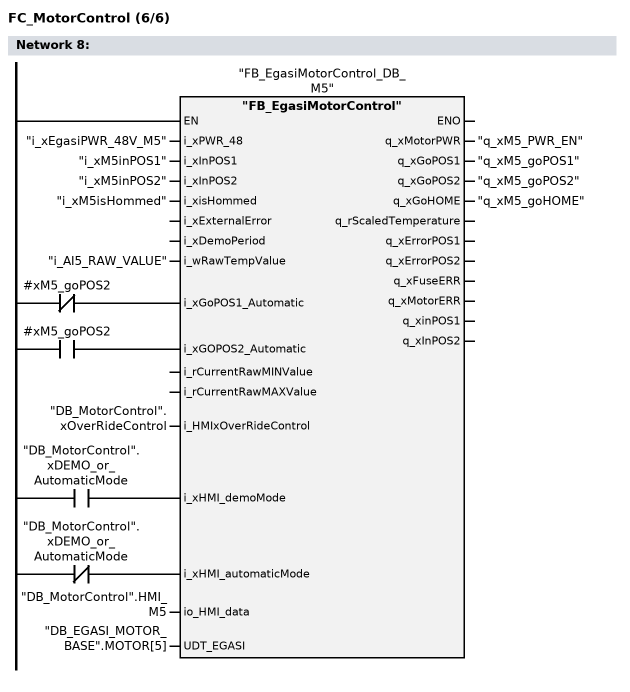
   RUNG wire#powerrail
      "FB_EgasiMotorControl_DB_M5"(i_xGoPOS1_Automatic := wire#w1, i_xGOPOS2_Automatic := wire#w2, i_xHMI_demoMode := wire#w3, i_xHMI_automaticMode := wire#w4, i_xPWR_48 := "i_xEgasiPWR_48V_M5", i_xInPOS1 := "i_xM5inPOS1", i_xInPOS2 := "i_xM5inPOS2", i_xisHommed := "i_xM5isHommed", i_xExternalError :=, i_xDemoPeriod :=, i_wRawTempValue := "i_AI5_RAW_VALUE", i_rCurrentRawMINValue :=, i_rCurrentRawMAXValue :=, i_HMIxOverRideControl := "DB_MotorControl".xOverRideControl, io_HMI_data := "DB_MotorControl".HMI_M5, UDT_EGASI := "DB_EGASI_MOTOR_BASE".MOTOR[5], q_xMotorPWR => "q_xM5_PWR_EN", q_xGoPOS1 => "q_xM5_goPOS1", q_xGoPOS2 => "q_xM5_goPOS2", q_xGoHOME => "q_xM5_goHOME", q_rScaledTemperature =>, q_xErrorPOS1 =>, q_xErrorPOS2 =>, q_xFuseERR =>, q_xMotorERR =>, q_xinPOS1 =>, q_xInPOS2 =>)
   END_RUNG
   RUNG wire#powerrail
      I_Contact( #xM5_goPOS2 )
   END_RUNG wire#w1
   RUNG wire#powerrail
      Contact( #xM5_goPOS2 )
   END_RUNG wire#w2
   RUNG wire#powerrail
      Contact( "DB_MotorControl".xDEMO_or_AutomaticMode )
   END_RUNG wire#w3
   RUNG wire#powerrail
      I_Contact( "DB_MotorControl".xDEMO_or_AutomaticMode )
   END_RUNG wire#w4
   // the same network as SCL:
   "FB_EgasiMotorControl_DB_M5"(i_xPWR_48 := "i_xEgasiPWR_48V_M5",   // "FB_EgasiMotorControl"
                           i_xInPOS1 := "i_xM5inPOS1",
                           i_xInPOS2 := "i_xM5inPOS2",
                           i_xisHommed := "i_xM5isHommed",
                           i_wRawTempValue := "i_AI5_RAW_VALUE",
                           i_xGoPOS1_Automatic := NOT #xM5_goPOS2,
                           i_xGOPOS2_Automatic := #xM5_goPOS2,
                           i_HMIxOverRideControl := "DB_MotorControl".xOverRideControl,
                           i_xHMI_demoMode := "DB_MotorControl".xDEMO_or_AutomaticMode,
                           i_xHMI_automaticMode := NOT "DB_MotorControl".xDEMO_or_AutomaticMode,
                           io_HMI_data := "DB_MotorControl".HMI_M5,
                           UDT_EGASI := "DB_EGASI_MOTOR_BASE".MOTOR[5],
                           q_xMotorPWR => "q_xM5_PWR_EN",
                           q_xGoPOS1 => "q_xM5_goPOS1",
                           q_xGoPOS2 => "q_xM5_goPOS2",
                           q_xGoHOME => "q_xM5_goHOME");
END_REGION
END_FUNCTION

FUNCTION "FC_PARTMANAGE" : Void   // FC12, LAD
{ S7_Optimized_Access := 'TRUE' }
VERSION : 0.1
   VAR_TEMP   // added for the SCL form of the ladder/FBD networks
      _w1 : Bool;
   END_VAR
BEGIN

REGION Network 2: COPY DATA FROM BASE TO DB for Cylinder control
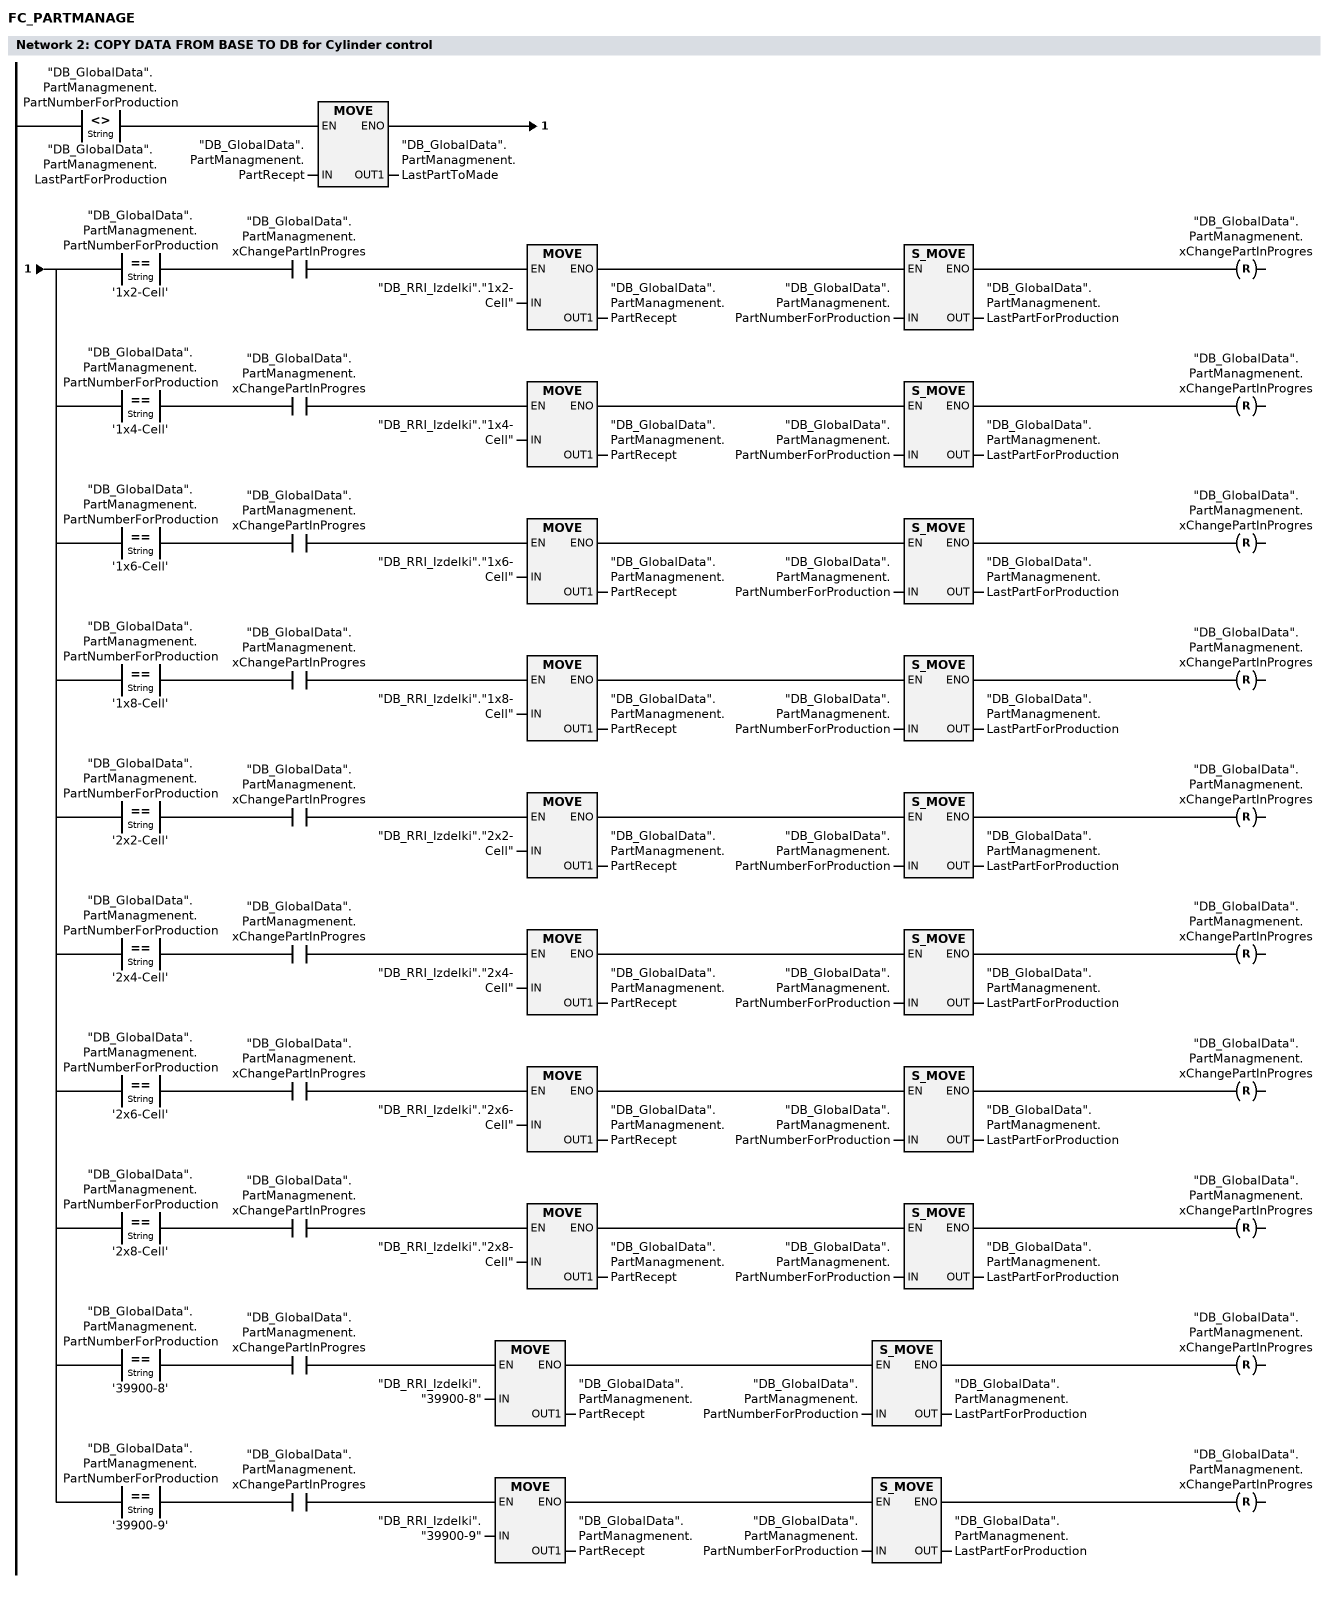
   RUNG wire#powerrail
      { S7_Templates := "SrcType := String" } NE_Contact(in1 := "DB_GlobalData".PartManagmenent.PartNumberForProduction, in2 := "DB_GlobalData".PartManagmenent.LastPartForProduction)
      Move(in := "DB_GlobalData".PartManagmenent.PartRecept, out1 => "DB_GlobalData".PartManagmenent.LastPartToMade)
      wire#w1
      { S7_Templates := "SrcType := String" } EQ_Contact(in1 := "DB_GlobalData".PartManagmenent.PartNumberForProduction, in2 := '1x2-Cell')
      Contact( "DB_GlobalData".PartManagmenent.xChangePartInProgres )
      Move(in := "DB_RRI_Izdelki"."1x2-Cell", out1 => "DB_GlobalData".PartManagmenent.PartRecept)
      S_Move(in := "DB_GlobalData".PartManagmenent.PartNumberForProduction, out => "DB_GlobalData".PartManagmenent.LastPartForProduction)
      R_Coil( "DB_GlobalData".PartManagmenent.xChangePartInProgres )
   END_RUNG
   RUNG wire#w1
      { S7_Templates := "SrcType := String" } EQ_Contact(in1 := "DB_GlobalData".PartManagmenent.PartNumberForProduction, in2 := '1x4-Cell')
      Contact( "DB_GlobalData".PartManagmenent.xChangePartInProgres )
      Move(in := "DB_RRI_Izdelki"."1x4-Cell", out1 => "DB_GlobalData".PartManagmenent.PartRecept)
      S_Move(in := "DB_GlobalData".PartManagmenent.PartNumberForProduction, out => "DB_GlobalData".PartManagmenent.LastPartForProduction)
      R_Coil( "DB_GlobalData".PartManagmenent.xChangePartInProgres )
   END_RUNG
   RUNG wire#w1
      { S7_Templates := "SrcType := String" } EQ_Contact(in1 := "DB_GlobalData".PartManagmenent.PartNumberForProduction, in2 := '1x6-Cell')
      Contact( "DB_GlobalData".PartManagmenent.xChangePartInProgres )
      Move(in := "DB_RRI_Izdelki"."1x6-Cell", out1 => "DB_GlobalData".PartManagmenent.PartRecept)
      S_Move(in := "DB_GlobalData".PartManagmenent.PartNumberForProduction, out => "DB_GlobalData".PartManagmenent.LastPartForProduction)
      R_Coil( "DB_GlobalData".PartManagmenent.xChangePartInProgres )
   END_RUNG
   RUNG wire#w1
      { S7_Templates := "SrcType := String" } EQ_Contact(in1 := "DB_GlobalData".PartManagmenent.PartNumberForProduction, in2 := '1x8-Cell')
      Contact( "DB_GlobalData".PartManagmenent.xChangePartInProgres )
      Move(in := "DB_RRI_Izdelki"."1x8-Cell", out1 => "DB_GlobalData".PartManagmenent.PartRecept)
      S_Move(in := "DB_GlobalData".PartManagmenent.PartNumberForProduction, out => "DB_GlobalData".PartManagmenent.LastPartForProduction)
      R_Coil( "DB_GlobalData".PartManagmenent.xChangePartInProgres )
   END_RUNG
   RUNG wire#w1
      { S7_Templates := "SrcType := String" } EQ_Contact(in1 := "DB_GlobalData".PartManagmenent.PartNumberForProduction, in2 := '2x2-Cell')
      Contact( "DB_GlobalData".PartManagmenent.xChangePartInProgres )
      Move(in := "DB_RRI_Izdelki"."2x2-Cell", out1 => "DB_GlobalData".PartManagmenent.PartRecept)
      S_Move(in := "DB_GlobalData".PartManagmenent.PartNumberForProduction, out => "DB_GlobalData".PartManagmenent.LastPartForProduction)
      R_Coil( "DB_GlobalData".PartManagmenent.xChangePartInProgres )
   END_RUNG
   RUNG wire#w1
      { S7_Templates := "SrcType := String" } EQ_Contact(in1 := "DB_GlobalData".PartManagmenent.PartNumberForProduction, in2 := '2x4-Cell')
      Contact( "DB_GlobalData".PartManagmenent.xChangePartInProgres )
      Move(in := "DB_RRI_Izdelki"."2x4-Cell", out1 => "DB_GlobalData".PartManagmenent.PartRecept)
      S_Move(in := "DB_GlobalData".PartManagmenent.PartNumberForProduction, out => "DB_GlobalData".PartManagmenent.LastPartForProduction)
      R_Coil( "DB_GlobalData".PartManagmenent.xChangePartInProgres )
   END_RUNG
   RUNG wire#w1
      { S7_Templates := "SrcType := String" } EQ_Contact(in1 := "DB_GlobalData".PartManagmenent.PartNumberForProduction, in2 := '2x6-Cell')
      Contact( "DB_GlobalData".PartManagmenent.xChangePartInProgres )
      Move(in := "DB_RRI_Izdelki"."2x6-Cell", out1 => "DB_GlobalData".PartManagmenent.PartRecept)
      S_Move(in := "DB_GlobalData".PartManagmenent.PartNumberForProduction, out => "DB_GlobalData".PartManagmenent.LastPartForProduction)
      R_Coil( "DB_GlobalData".PartManagmenent.xChangePartInProgres )
   END_RUNG
   RUNG wire#w1
      { S7_Templates := "SrcType := String" } EQ_Contact(in1 := "DB_GlobalData".PartManagmenent.PartNumberForProduction, in2 := '2x8-Cell')
      Contact( "DB_GlobalData".PartManagmenent.xChangePartInProgres )
      Move(in := "DB_RRI_Izdelki"."2x8-Cell", out1 => "DB_GlobalData".PartManagmenent.PartRecept)
      S_Move(in := "DB_GlobalData".PartManagmenent.PartNumberForProduction, out => "DB_GlobalData".PartManagmenent.LastPartForProduction)
      R_Coil( "DB_GlobalData".PartManagmenent.xChangePartInProgres )
   END_RUNG
   RUNG wire#w1
      { S7_Templates := "SrcType := String" } EQ_Contact(in1 := "DB_GlobalData".PartManagmenent.PartNumberForProduction, in2 := '39900-8')
      Contact( "DB_GlobalData".PartManagmenent.xChangePartInProgres )
      Move(in := "DB_RRI_Izdelki"."39900-8", out1 => "DB_GlobalData".PartManagmenent.PartRecept)
      S_Move(in := "DB_GlobalData".PartManagmenent.PartNumberForProduction, out => "DB_GlobalData".PartManagmenent.LastPartForProduction)
      R_Coil( "DB_GlobalData".PartManagmenent.xChangePartInProgres )
   END_RUNG
   RUNG wire#w1
      { S7_Templates := "SrcType := String" } EQ_Contact(in1 := "DB_GlobalData".PartManagmenent.PartNumberForProduction, in2 := '39900-9')
      Contact( "DB_GlobalData".PartManagmenent.xChangePartInProgres )
      Move(in := "DB_RRI_Izdelki"."39900-9", out1 => "DB_GlobalData".PartManagmenent.PartRecept)
      S_Move(in := "DB_GlobalData".PartManagmenent.PartNumberForProduction, out => "DB_GlobalData".PartManagmenent.LastPartForProduction)
      R_Coil( "DB_GlobalData".PartManagmenent.xChangePartInProgres )
   END_RUNG
   // the same network as SCL:
   #_w1 := "DB_GlobalData".PartManagmenent.PartNumberForProduction <> "DB_GlobalData".PartManagmenent.LastPartForProduction;
   IF #_w1 THEN
       "DB_GlobalData".PartManagmenent.LastPartToMade := "DB_GlobalData".PartManagmenent.PartRecept;
   END_IF;
   IF #_w1 AND ("DB_GlobalData".PartManagmenent.PartNumberForProduction = '1x2-Cell') AND "DB_GlobalData".PartManagmenent.xChangePartInProgres THEN
       "DB_GlobalData".PartManagmenent.PartRecept := "DB_RRI_Izdelki"."1x2-Cell";
       "DB_GlobalData".PartManagmenent.LastPartForProduction := "DB_GlobalData".PartManagmenent.PartNumberForProduction;
       "DB_GlobalData".PartManagmenent.xChangePartInProgres := FALSE;
   END_IF;
   IF #_w1 AND ("DB_GlobalData".PartManagmenent.PartNumberForProduction = '1x4-Cell') AND "DB_GlobalData".PartManagmenent.xChangePartInProgres THEN
       "DB_GlobalData".PartManagmenent.PartRecept := "DB_RRI_Izdelki"."1x4-Cell";
       "DB_GlobalData".PartManagmenent.LastPartForProduction := "DB_GlobalData".PartManagmenent.PartNumberForProduction;
       "DB_GlobalData".PartManagmenent.xChangePartInProgres := FALSE;
   END_IF;
   IF #_w1 AND ("DB_GlobalData".PartManagmenent.PartNumberForProduction = '1x6-Cell') AND "DB_GlobalData".PartManagmenent.xChangePartInProgres THEN
       "DB_GlobalData".PartManagmenent.PartRecept := "DB_RRI_Izdelki"."1x6-Cell";
       "DB_GlobalData".PartManagmenent.LastPartForProduction := "DB_GlobalData".PartManagmenent.PartNumberForProduction;
       "DB_GlobalData".PartManagmenent.xChangePartInProgres := FALSE;
   END_IF;
   IF #_w1 AND ("DB_GlobalData".PartManagmenent.PartNumberForProduction = '1x8-Cell') AND "DB_GlobalData".PartManagmenent.xChangePartInProgres THEN
       "DB_GlobalData".PartManagmenent.PartRecept := "DB_RRI_Izdelki"."1x8-Cell";
       "DB_GlobalData".PartManagmenent.LastPartForProduction := "DB_GlobalData".PartManagmenent.PartNumberForProduction;
       "DB_GlobalData".PartManagmenent.xChangePartInProgres := FALSE;
   END_IF;
   IF #_w1 AND ("DB_GlobalData".PartManagmenent.PartNumberForProduction = '2x2-Cell') AND "DB_GlobalData".PartManagmenent.xChangePartInProgres THEN
       "DB_GlobalData".PartManagmenent.PartRecept := "DB_RRI_Izdelki"."2x2-Cell";
       "DB_GlobalData".PartManagmenent.LastPartForProduction := "DB_GlobalData".PartManagmenent.PartNumberForProduction;
       "DB_GlobalData".PartManagmenent.xChangePartInProgres := FALSE;
   END_IF;
   IF #_w1 AND ("DB_GlobalData".PartManagmenent.PartNumberForProduction = '2x4-Cell') AND "DB_GlobalData".PartManagmenent.xChangePartInProgres THEN
       "DB_GlobalData".PartManagmenent.PartRecept := "DB_RRI_Izdelki"."2x4-Cell";
       "DB_GlobalData".PartManagmenent.LastPartForProduction := "DB_GlobalData".PartManagmenent.PartNumberForProduction;
       "DB_GlobalData".PartManagmenent.xChangePartInProgres := FALSE;
   END_IF;
   IF #_w1 AND ("DB_GlobalData".PartManagmenent.PartNumberForProduction = '2x6-Cell') AND "DB_GlobalData".PartManagmenent.xChangePartInProgres THEN
       "DB_GlobalData".PartManagmenent.PartRecept := "DB_RRI_Izdelki"."2x6-Cell";
       "DB_GlobalData".PartManagmenent.LastPartForProduction := "DB_GlobalData".PartManagmenent.PartNumberForProduction;
       "DB_GlobalData".PartManagmenent.xChangePartInProgres := FALSE;
   END_IF;
   IF #_w1 AND ("DB_GlobalData".PartManagmenent.PartNumberForProduction = '2x8-Cell') AND "DB_GlobalData".PartManagmenent.xChangePartInProgres THEN
       "DB_GlobalData".PartManagmenent.PartRecept := "DB_RRI_Izdelki"."2x8-Cell";
       "DB_GlobalData".PartManagmenent.LastPartForProduction := "DB_GlobalData".PartManagmenent.PartNumberForProduction;
       "DB_GlobalData".PartManagmenent.xChangePartInProgres := FALSE;
   END_IF;
   IF #_w1 AND ("DB_GlobalData".PartManagmenent.PartNumberForProduction = '39900-8') AND "DB_GlobalData".PartManagmenent.xChangePartInProgres THEN
       "DB_GlobalData".PartManagmenent.PartRecept := "DB_RRI_Izdelki"."39900-8";
       "DB_GlobalData".PartManagmenent.LastPartForProduction := "DB_GlobalData".PartManagmenent.PartNumberForProduction;
       "DB_GlobalData".PartManagmenent.xChangePartInProgres := FALSE;
   END_IF;
   IF #_w1 AND ("DB_GlobalData".PartManagmenent.PartNumberForProduction = '39900-9') AND "DB_GlobalData".PartManagmenent.xChangePartInProgres THEN
       "DB_GlobalData".PartManagmenent.PartRecept := "DB_RRI_Izdelki"."39900-9";
       "DB_GlobalData".PartManagmenent.LastPartForProduction := "DB_GlobalData".PartManagmenent.PartNumberForProduction;
       "DB_GlobalData".PartManagmenent.xChangePartInProgres := FALSE;
   END_IF;
END_REGION

REGION Network 3 (SCL)
   // HMI read data
   // 
   IF ("DB_DATAFORCOMMUNICATION".iHMIpartNumber <>"DB_DATAFORCOMMUNICATION".iHmiLastPartNumber) AND
       "DB_GlobalData".PartManagmenent.Trenutni_pomik = 0 THEN
       //read part number
       CASE "DB_DATAFORCOMMUNICATION".iHMIpartNumber OF
           12:
               "DB_GlobalData".PartManagmenent.PartNumberForProduction := '1x2-Cell';
           14:
               "DB_GlobalData".PartManagmenent.PartNumberForProduction := '1x4-Cell';
           16:
               "DB_GlobalData".PartManagmenent.PartNumberForProduction := '1x6-Cell';
           18:
               "DB_GlobalData".PartManagmenent.PartNumberForProduction := '1x8-Cell';
           22:
               "DB_GlobalData".PartManagmenent.PartNumberForProduction := '2x2-Cell';
           24:
               "DB_GlobalData".PartManagmenent.PartNumberForProduction := '2x4-Cell';
           26:
               "DB_GlobalData".PartManagmenent.PartNumberForProduction := '2x6-Cell';
           28:
               "DB_GlobalData".PartManagmenent.PartNumberForProduction := '2x8-Cell';
           ELSE
               ;
               ;
       END_CASE;

       "DB_DATAFORCOMMUNICATION".iHmiLastPartNumber := "DB_DATAFORCOMMUNICATION".iHMIpartNumber;
   END_IF;
END_REGION

REGION Network 4: HMI read data
END_REGION
END_FUNCTION

FUNCTION "GetMotorOuput" : Void   // FC14, LAD
{ S7_Optimized_Access := 'TRUE' }
VERSION : 0.1
   VAR_INPUT
      recept_id : Int;
      motorNO : Int;
      feed_pos : Int;
   END_VAR
   VAR_OUTPUT
      GetMotorOutput : Bool;
   END_VAR
   VAR_IN_OUT
      Recipe_1x2 : "RRI_izdelki";
      Recipe_1x4 : "RRI_izdelki";
      Recipe_1x6 : "RRI_izdelki";
      Recipe_1x8 : "RRI_izdelki";
      Recipe_2x2 : "RRI_izdelki";
      Recipe_2x4 : "RRI_izdelki";
      Recipe_2x6 : "RRI_izdelki";
      Recipe_2x8 : "RRI_izdelki";
   END_VAR
BEGIN

REGION Network 2 (SCL)
   CASE #recept_id OF
       12:
           CASE #motorNO OF
               1:
                   #GetMotorOutput := #Recipe_1x2.NazivniPodatki.CILINDRI.MOTOR1[#feed_pos];
               2:
                   #GetMotorOutput := #Recipe_1x2.NazivniPodatki.CILINDRI.MOTOR2[#feed_pos];
               3:
                   #GetMotorOutput := #Recipe_1x2.NazivniPodatki.CILINDRI.MOTOR3[#feed_pos];
               4:
                   #GetMotorOutput := #Recipe_1x2.NazivniPodatki.CILINDRI.MOTOR4[#feed_pos];
               5:
                   #GetMotorOutput := #Recipe_1x2.NazivniPodatki.CILINDRI.MOTOR5[#feed_pos];
           END_CASE;

       14:
           CASE #motorNO OF
               1:
                   #GetMotorOutput := #Recipe_1x4.NazivniPodatki.CILINDRI.MOTOR1[#feed_pos];
               2:
                   #GetMotorOutput := #Recipe_1x4.NazivniPodatki.CILINDRI.MOTOR2[#feed_pos];
               3:
                   #GetMotorOutput := #Recipe_1x4.NazivniPodatki.CILINDRI.MOTOR3[#feed_pos];
               4:
                   #GetMotorOutput := #Recipe_1x4.NazivniPodatki.CILINDRI.MOTOR4[#feed_pos];
               5:
                   #GetMotorOutput := #Recipe_1x4.NazivniPodatki.CILINDRI.MOTOR5[#feed_pos];
           END_CASE;

       16:
           CASE #motorNO OF
               1:
                   #GetMotorOutput := #Recipe_1x6.NazivniPodatki.CILINDRI.MOTOR1[#feed_pos];
               2:
                   #GetMotorOutput := #Recipe_1x6.NazivniPodatki.CILINDRI.MOTOR2[#feed_pos];
               3:
                   #GetMotorOutput := #Recipe_1x6.NazivniPodatki.CILINDRI.MOTOR3[#feed_pos];
               4:
                   #GetMotorOutput := #Recipe_1x6.NazivniPodatki.CILINDRI.MOTOR4[#feed_pos];
               5:
                   #GetMotorOutput := #Recipe_1x6.NazivniPodatki.CILINDRI.MOTOR5[#feed_pos];
           END_CASE;

       18:
           CASE #motorNO OF
               1:
                   #GetMotorOutput := #Recipe_1x8.NazivniPodatki.CILINDRI.MOTOR1[#feed_pos];
               2:
                   #GetMotorOutput := #Recipe_1x8.NazivniPodatki.CILINDRI.MOTOR2[#feed_pos];
               3:
                   #GetMotorOutput := #Recipe_1x8.NazivniPodatki.CILINDRI.MOTOR3[#feed_pos];
               4:
                   #GetMotorOutput := #Recipe_1x8.NazivniPodatki.CILINDRI.MOTOR4[#feed_pos];
               5:
                   #GetMotorOutput := #Recipe_1x8.NazivniPodatki.CILINDRI.MOTOR5[#feed_pos];
           END_CASE;

       22:
           CASE #motorNO OF
               1:
                   #GetMotorOutput := #Recipe_2x2.NazivniPodatki.CILINDRI.MOTOR1[#feed_pos];
               2:
                   #GetMotorOutput := #Recipe_2x2.NazivniPodatki.CILINDRI.MOTOR2[#feed_pos];
               3:
                   #GetMotorOutput := #Recipe_2x2.NazivniPodatki.CILINDRI.MOTOR3[#feed_pos];
               4:
                   #GetMotorOutput := #Recipe_2x2.NazivniPodatki.CILINDRI.MOTOR4[#feed_pos];
               5:
                   #GetMotorOutput := #Recipe_2x2.NazivniPodatki.CILINDRI.MOTOR5[#feed_pos];
           END_CASE;

       24:
           CASE #motorNO OF
               1:
                   #GetMotorOutput := #Recipe_2x4.NazivniPodatki.CILINDRI.MOTOR1[#feed_pos];
               2:
                   #GetMotorOutput := #Recipe_2x4.NazivniPodatki.CILINDRI.MOTOR2[#feed_pos];
               3:
                   #GetMotorOutput := #Recipe_2x4.NazivniPodatki.CILINDRI.MOTOR3[#feed_pos];
               4:
                   #GetMotorOutput := #Recipe_2x4.NazivniPodatki.CILINDRI.MOTOR4[#feed_pos];
               5:
                   #GetMotorOutput := #Recipe_2x4.NazivniPodatki.CILINDRI.MOTOR5[#feed_pos];
           END_CASE;

       26:
           CASE #motorNO OF
               1:
                   #GetMotorOutput := #Recipe_2x6.NazivniPodatki.CILINDRI.MOTOR1[#feed_pos];
               2:
                   #GetMotorOutput := #Recipe_2x6.NazivniPodatki.CILINDRI.MOTOR2[#feed_pos];
               3:
                   #GetMotorOutput := #Recipe_2x6.NazivniPodatki.CILINDRI.MOTOR3[#feed_pos];
               4:
                   #GetMotorOutput := #Recipe_2x6.NazivniPodatki.CILINDRI.MOTOR4[#feed_pos];
               5:
                   #GetMotorOutput := #Recipe_2x6.NazivniPodatki.CILINDRI.MOTOR5[#feed_pos];
           END_CASE;

       28:
           CASE #motorNO OF
               1:
                   #GetMotorOutput := #Recipe_2x8.NazivniPodatki.CILINDRI.MOTOR1[#feed_pos];
               2:
                   #GetMotorOutput := #Recipe_2x8.NazivniPodatki.CILINDRI.MOTOR2[#feed_pos];
               3:
                   #GetMotorOutput := #Recipe_2x8.NazivniPodatki.CILINDRI.MOTOR3[#feed_pos];
               4:
                   #GetMotorOutput := #Recipe_2x8.NazivniPodatki.CILINDRI.MOTOR4[#feed_pos];
               5:
                   #GetMotorOutput := #Recipe_2x8.NazivniPodatki.CILINDRI.MOTOR5[#feed_pos];
           END_CASE;

       ELSE
           #GetMotorOutput := FALSE; // default off
   END_CASE;
END_REGION
END_FUNCTION

FUNCTION "FC_GetMaxFeeds" : Void   // FC15, LAD
{ S7_Optimized_Access := 'TRUE' }
VERSION : 0.1
   VAR_INPUT
      recept_id : Int;
   END_VAR
   VAR_OUTPUT
      GetMaxFeeds : Int;
   END_VAR
   VAR_IN_OUT
      Recipe_2x2 : "RRI_izdelki";
      Recipe_2x4 : "RRI_izdelki";
      Recipe_2x6 : "RRI_izdelki";
      Recipe_2x8 : "RRI_izdelki";
      Recipe_1x2 : "RRI_izdelki";
      Recipe_1x4 : "RRI_izdelki";
      Recipe_1x6 : "RRI_izdelki";
      Recipe_1x8 : "RRI_izdelki";
   END_VAR
BEGIN

REGION Network 2 (SCL)
   CASE #recept_id OF
       12:
           #GetMaxFeeds := #Recipe_2x2.NazivniPodatki.st_pomikov;   // st_pomikov = max index (1)
       24:
           #GetMaxFeeds := #Recipe_2x4.NazivniPodatki.st_pomikov;   // (3)
       26:
           #GetMaxFeeds := #Recipe_2x6.NazivniPodatki.st_pomikov;   // (5)
       28:
           #GetMaxFeeds := #Recipe_2x8.NazivniPodatki.st_pomikov;   // (7)
       14:
           #GetMaxFeeds := #Recipe_1x4.NazivniPodatki.st_pomikov;   // etc.
       16:
           #GetMaxFeeds := #Recipe_1x6.NazivniPodatki.st_pomikov;
       18:
           #GetMaxFeeds := #Recipe_1x2.NazivniPodatki.st_pomikov;
       12:
           #GetMaxFeeds := #Recipe_1x2.NazivniPodatki.st_pomikov;
       ELSE
           #GetMaxFeeds := 0;
   END_CASE;
END_REGION
END_FUNCTION

ORGANIZATION_BLOCK "Main"   // OB1, LAD, ProgramCycle
TITLE = "Main Program Sweep (Cycle)"
{ S7_Optimized_Access := 'TRUE' }
VERSION : 0.1
   VAR_INPUT
      Initial_Call : Bool;   // Initial call of this OB
      Remanence : Bool;   // =True, if remanent data are available
   END_VAR
   VAR_TEMP   // added for the SCL form of the ladder/FBD networks
      _w1 : Bool;
      _w2 : Bool;
   END_VAR
BEGIN

REGION Network 1
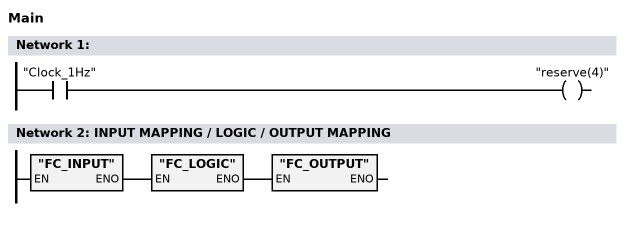
   RUNG wire#powerrail
      Contact( "Clock_1Hz" )
      Coil( "reserve(4)" )
   END_RUNG
   // the same network as SCL:
   "reserve(4)" := "Clock_1Hz";
END_REGION

REGION Network 2: INPUT MAPPING / LOGIC / OUTPUT MAPPING
   RUNG wire#powerrail
      "FC_INPUT"()
      "FC_LOGIC"()
      "FC_OUTPUT"()
   END_RUNG
   // the same network as SCL:
   "FC_INPUT"(ENO => #_w1);
   "FC_LOGIC"(EN := #_w1, ENO => #_w2);
   IF #_w2 THEN "FC_OUTPUT"(); END_IF;
END_REGION
END_ORGANIZATION_BLOCK

// folder: AKD

FUNCTION_BLOCK "FB_AKD"   // FB11, LAD
{ S7_Optimized_Access := 'TRUE' }
VERSION : 0.1
   VAR_INPUT
      bServoEnable : Bool;
      iNastavitevHitrosti : Int;
      dNastavitevPozicije : DInt;
      bPogojiZaVKLOP : Bool;
      iAKD : "AKD_TO_SIEMENS";
      ResetNapake : Bool;
      iStPrograma : Word;
   END_VAR
   VAR_OUTPUT
      oAKD : "SIEMENS_TO_AKD";
      AKDcurrPos : DInt;
      o_BerrStatus : Byte;
      rAKDpos : Real;
      xDriveIsStoped : Bool;
      q_xStartHomming : Bool;
      q_xisHommed : Bool;
      q_xerrNoInTolleranceRange : Bool;
   END_VAR
   VAR_IN_OUT
      iStartHoming : Bool;
      bServoGo : Bool;
   END_VAR
   VAR RETAIN
      TIMER_ON : Array[0..5] of TON_TIME;
   END_VAR
   VAR
      diHitrost : Real;
      dwHitrostRez : Real;
      ServoHommed : Bool;
   END_VAR
   VAR RETAIN
      merker : Array[0..1] of Bool;
   END_VAR
   VAR
      OmogociHome : Bool;
      Varnost : Bool;
      M_varnost : Bool;
      varnostN : Bool;
      TON_fault : TON_TIME;
   END_VAR
   VAR RETAIN
      _xServoGoP : Bool;
      _rCurrntPosition : Real;
      _xServoGoN : Bool;
      _xLastPosition : Real;
   END_VAR
   VAR
      IEC_Timer_0_Instance : TP_TIME;
      R_TRIG_Instance_Home : R_TRIG;
   END_VAR
   VAR RETAIN
      "p_trig-HomePosSet" : Bool;
      "P-trig" : Bool;
      MDI_STATUS : Int;
   END_VAR
   VAR
      statis_target_pos_reach : Bool;
      _errorNotInToleranceRange : Bool;
   END_VAR
   VAR CONSTANT
      AXES_START_MOVING : Int := 10;
      TARGET_POS_REACH : Int := 20;
      RESET_SERVO_GO : Int := 30;
   END_VAR
   VAR_TEMP   // added for the SCL form of the ladder/FBD networks
      _w1 : Bool;
      _w2 : Bool;
      _w3 : Bool;
      _w4 : Bool;
   END_VAR
BEGIN

REGION Network 1: Bool
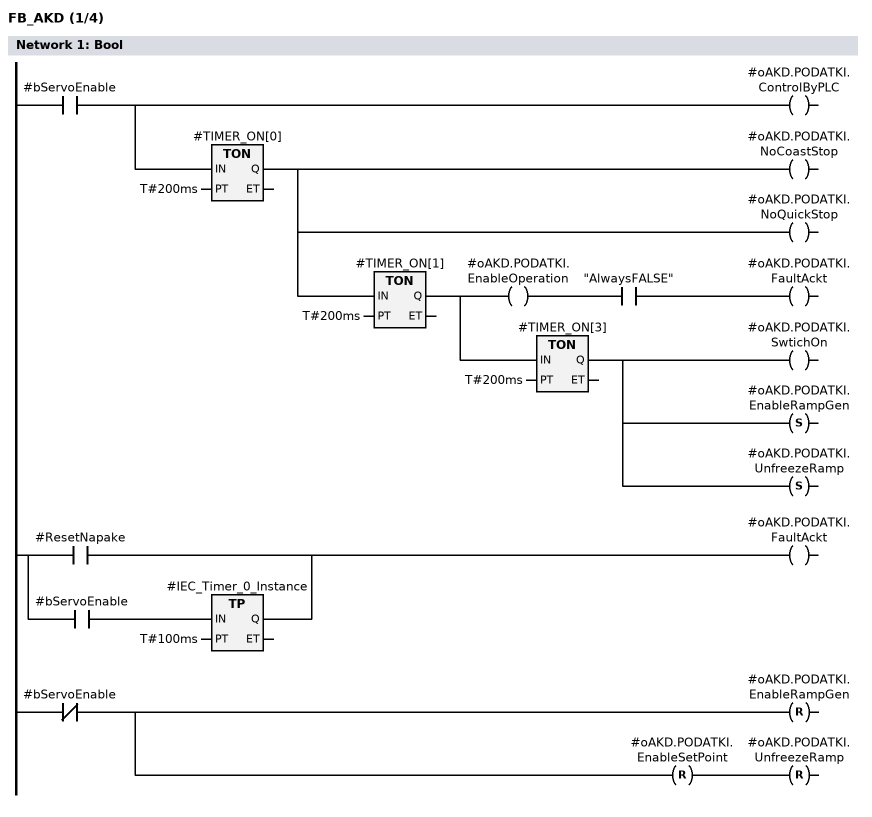
   #oAKD.PODATKI.ControlByPLC := #bServoEnable;
   #TIMER_ON[0].TON(IN := #bServoEnable, PT := T#200ms);
   #oAKD.PODATKI.NoCoastStop := #TIMER_ON[0].Q;
   #oAKD.PODATKI.NoQuickStop := #TIMER_ON[0].Q;
   #TIMER_ON[1].TON(IN := #TIMER_ON[0].Q, PT := T#200ms);
   #oAKD.PODATKI.EnableOperation := #TIMER_ON[1].Q;
   #oAKD.PODATKI.FaultAckt := #TIMER_ON[1].Q AND "AlwaysFALSE";
   #TIMER_ON[3].TON(IN := #TIMER_ON[1].Q, PT := T#200ms);
   #oAKD.PODATKI.SwtichOn := #TIMER_ON[3].Q;
   IF #TIMER_ON[3].Q THEN
       #oAKD.PODATKI.EnableRampGen := TRUE;
       #oAKD.PODATKI.UnfreezeRamp := TRUE;
   END_IF;
   #IEC_Timer_0_Instance(IN := #bServoEnable, PT := T#100ms);   // TP
   #oAKD.PODATKI.FaultAckt := #ResetNapake OR #IEC_Timer_0_Instance.Q;
   IF NOT #bServoEnable THEN
       #oAKD.PODATKI.EnableRampGen := FALSE;
       #oAKD.PODATKI.EnableSetPoint := FALSE;
       #oAKD.PODATKI.UnfreezeRamp := FALSE;
   END_IF;
END_REGION

REGION Network 2: Turn on MDI - manual data inpuit - start task on AKD
   // Requeremnts
   // - S4
   // - mode in position mode (yes)
   // - standard telegram 9 (set at profinet configuration)
   // - axis hommed (homeposset)
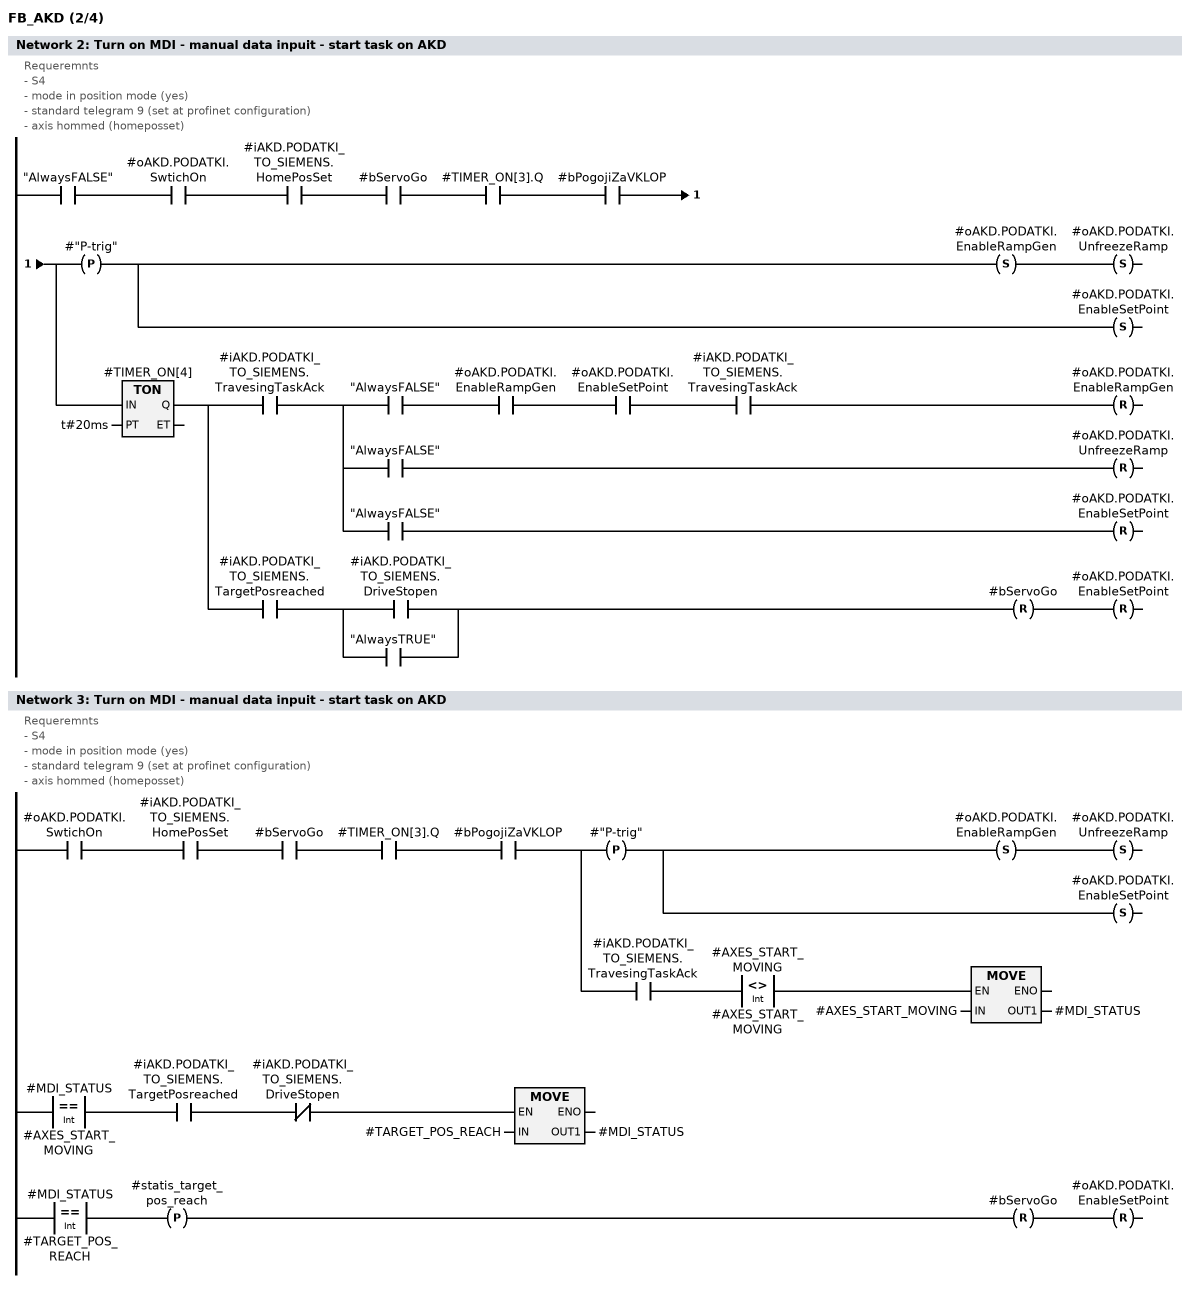
   #_w1 := "AlwaysFALSE" AND #oAKD.PODATKI.SwtichOn AND #iAKD.PODATKI_TO_SIEMENS.HomePosSet AND #bServoGo AND #TIMER_ON[3].Q AND #bPogojiZaVKLOP;
   #_w2 := #_w1 AND NOT #"P-trig";   // rising edge
   #"P-trig" := #_w1;
   IF #_w2 THEN
       #oAKD.PODATKI.EnableRampGen := TRUE;
       #oAKD.PODATKI.UnfreezeRamp := TRUE;
       #oAKD.PODATKI.EnableSetPoint := TRUE;
   END_IF;
   #TIMER_ON[4].TON(IN := #_w1, PT := t#20ms);
   #_w3 := #TIMER_ON[4].Q AND #iAKD.PODATKI_TO_SIEMENS.TravesingTaskAck;
   IF #_w3 AND "AlwaysFALSE" AND #oAKD.PODATKI.EnableRampGen AND #oAKD.PODATKI.EnableSetPoint AND #iAKD.PODATKI_TO_SIEMENS.TravesingTaskAck THEN
       #oAKD.PODATKI.EnableRampGen := FALSE;
   END_IF;
   IF #_w3 AND "AlwaysFALSE" THEN
       #oAKD.PODATKI.UnfreezeRamp := FALSE;
       #oAKD.PODATKI.EnableSetPoint := FALSE;
   END_IF;
   IF #TIMER_ON[4].Q AND #iAKD.PODATKI_TO_SIEMENS.TargetPosreached AND (#iAKD.PODATKI_TO_SIEMENS.DriveStopen OR "AlwaysTRUE") THEN
       #bServoGo := FALSE;
       #oAKD.PODATKI.EnableSetPoint := FALSE;
   END_IF;
END_REGION

REGION Network 3: Turn on MDI - manual data inpuit - start task on AKD
   // Requeremnts
   // - S4
   // - mode in position mode (yes)
   // - standard telegram 9 (set at profinet configuration)
   // - axis hommed (homeposset)
   RUNG wire#powerrail
      Contact( #oAKD.PODATKI.SwtichOn )
      Contact( #iAKD.PODATKI_TO_SIEMENS.HomePosSet )
      Contact( #bServoGo )
      Contact( #TIMER_ON[3].Q )
      Contact( #bPogojiZaVKLOP )
      wire#w1
      P_Trig( #"P-trig" )
      wire#w2
      S_Coil( #oAKD.PODATKI.EnableRampGen )
      S_Coil( #oAKD.PODATKI.UnfreezeRamp )
   END_RUNG
   RUNG wire#w2
      S_Coil( #oAKD.PODATKI.EnableSetPoint )
   END_RUNG
   RUNG wire#w1
      Contact( #iAKD.PODATKI_TO_SIEMENS.TravesingTaskAck )
      { S7_Templates := "SrcType := Int" } NE_Contact(in1 := #AXES_START_MOVING, in2 := #AXES_START_MOVING)
      Move(in := #AXES_START_MOVING, out1 => #MDI_STATUS)
   END_RUNG
   RUNG wire#powerrail
      { S7_Templates := "SrcType := Int" } EQ_Contact(in1 := #MDI_STATUS, in2 := #AXES_START_MOVING)
      Contact( #iAKD.PODATKI_TO_SIEMENS.TargetPosreached )
      I_Contact( #iAKD.PODATKI_TO_SIEMENS.DriveStopen )
      Move(in := #TARGET_POS_REACH, out1 => #MDI_STATUS)
   END_RUNG
   RUNG wire#powerrail
      { S7_Templates := "SrcType := Int" } EQ_Contact(in1 := #MDI_STATUS, in2 := #TARGET_POS_REACH)
      P_Trig( #statis_target_pos_reach )
      R_Coil( #bServoGo )
      R_Coil( #oAKD.PODATKI.EnableSetPoint )
   END_RUNG
   // the same network as SCL:
   #_w1 := #oAKD.PODATKI.SwtichOn AND #iAKD.PODATKI_TO_SIEMENS.HomePosSet AND #bServoGo AND #TIMER_ON[3].Q AND #bPogojiZaVKLOP;
   #_w2 := #_w1 AND NOT #"P-trig";   // rising edge
   #"P-trig" := #_w1;
   IF #_w2 THEN
       #oAKD.PODATKI.EnableRampGen := TRUE;
       #oAKD.PODATKI.UnfreezeRamp := TRUE;
       #oAKD.PODATKI.EnableSetPoint := TRUE;
   END_IF;
   IF #_w1 AND #iAKD.PODATKI_TO_SIEMENS.TravesingTaskAck AND (#AXES_START_MOVING <> #AXES_START_MOVING) THEN
       #MDI_STATUS := #AXES_START_MOVING;
   END_IF;
   IF (#MDI_STATUS = #AXES_START_MOVING) AND #iAKD.PODATKI_TO_SIEMENS.TargetPosreached AND NOT #iAKD.PODATKI_TO_SIEMENS.DriveStopen THEN
       #MDI_STATUS := #TARGET_POS_REACH;
   END_IF;
   #_w3 := #MDI_STATUS = #TARGET_POS_REACH;
   #_w4 := #_w3 AND NOT #statis_target_pos_reach;   // rising edge
   #statis_target_pos_reach := #_w3;
   IF #_w4 THEN
       #bServoGo := FALSE;
       #oAKD.PODATKI.EnableSetPoint := FALSE;
   END_IF;
END_REGION

REGION Network 4